REGION Network 108
   RUNG wire#powerrail
      Move(in := "Carrier_05_SDCFaultCode", out1 => "DB_SDC_EMS_TA".EMS[05].TA[1].FAULT)
      wire#w1
      Move(in := "Carrier_05_SDCFaultCode", out1 => "EMS".Carrier[05].SDC_IN.CarrierDriveFaults)
   END_RUNG
   RUNG wire#powerrail
      Contact( "IndiconTempDebugON" )
   END_RUNG wire#w1
   // the same network as SCL:
   "DB_SDC_EMS_TA".EMS[05].TA[1].FAULT := "Carrier_05_SDCFaultCode";
   IF TRUE OR "IndiconTempDebugON" THEN
       "EMS".Carrier[05].SDC_IN.CarrierDriveFaults := "Carrier_05_SDCFaultCode";
   END_IF;
END_REGION

REGION Network 109
   RUNG wire#powerrail
      Move(in := "Carrier_05_CarrierDriveAlarm", out1 => "DB_SDC_EMS_TA".EMS[05].TA[1].ALARM)
      wire#w1
      Move(in := "Carrier_05_CarrierDriveAlarm", out1 => "EMS".Carrier[05].SDC_IN.CarrierDriveAlarms)
   END_RUNG
   RUNG wire#powerrail
      Contact( "IndiconTempDebugON" )
   END_RUNG wire#w1
   // the same network as SCL:
   "DB_SDC_EMS_TA".EMS[05].TA[1].ALARM := "Carrier_05_CarrierDriveAlarm";
   IF TRUE OR "IndiconTempDebugON" THEN
       "EMS".Carrier[05].SDC_IN.CarrierDriveAlarms := "Carrier_05_CarrierDriveAlarm";
   END_IF;
END_REGION

REGION Network 110
   RUNG wire#powerrail
      Move(in := "Carrier_05_SDCFaultCode", out1 => "DB101_DB_SDC_FAULTS".Carrier_Fault[05])
      wire#w1
      Move(in := "Carrier_05_SDCFaultCode", out1 => "EMS".Carrier[05].SDC_IN.CarrierFaults)
   END_RUNG
   RUNG wire#powerrail
      Contact( "IndiconTempDebugON" )
   END_RUNG wire#w1
   // the same network as SCL:
   "DB101_DB_SDC_FAULTS".Carrier_Fault[05] := "Carrier_05_SDCFaultCode";
   IF TRUE OR "IndiconTempDebugON" THEN
       "EMS".Carrier[05].SDC_IN.CarrierFaults := "Carrier_05_SDCFaultCode";
   END_IF;
END_REGION

REGION Network 111
   RUNG wire#powerrail
      Contact( "Carrier_05_Status.5" )
      Coil( "EMS".Carrier[05].SDC_IN.RunningFWD )
   END_RUNG
   // the same network as SCL:
   "EMS".Carrier[05].SDC_IN.RunningFWD := "Carrier_05_Status.5";
END_REGION

REGION Network 112
   RUNG wire#powerrail
      Contact( "Carrier_05_Status.6" )
      Coil( "EMS".Carrier[05].SDC_IN.RunningREV )
   END_RUNG
   // the same network as SCL:
   "EMS".Carrier[05].SDC_IN.RunningREV := "Carrier_05_Status.6";
END_REGION

REGION Network 113
   RUNG wire#powerrail
      Contact( "Carrier_05_Status.7" )
      Coil( "EMS".Carrier[05].SDC_IN.IR_Remote_9_Pressed )
   END_RUNG
   // the same network as SCL:
   "EMS".Carrier[05].SDC_IN.IR_Remote_9_Pressed := "Carrier_05_Status.7";
END_REGION

REGION Network 114
   RUNG wire#powerrail
      I_Contact( "Carrier_05_Status.5" )
      I_Contact( "Carrier_05_Status.6" )
      Coil( "EMS".Carrier[05].SDC_IN.Stopped )
   END_RUNG
   // the same network as SCL:
   "EMS".Carrier[05].SDC_IN.Stopped := NOT "Carrier_05_Status.5" AND NOT "Carrier_05_Status.6";
END_REGION

REGION Network 115
   RUNG wire#powerrail
      Contact( "Carrier_05_Status.4" )
      Coil( "EMS".Carrier[05].SDC_IN.ProductionHoldPB_Status )
   END_RUNG
   // the same network as SCL:
   "EMS".Carrier[05].SDC_IN.ProductionHoldPB_Status := "Carrier_05_Status.4";
END_REGION

REGION Network 116
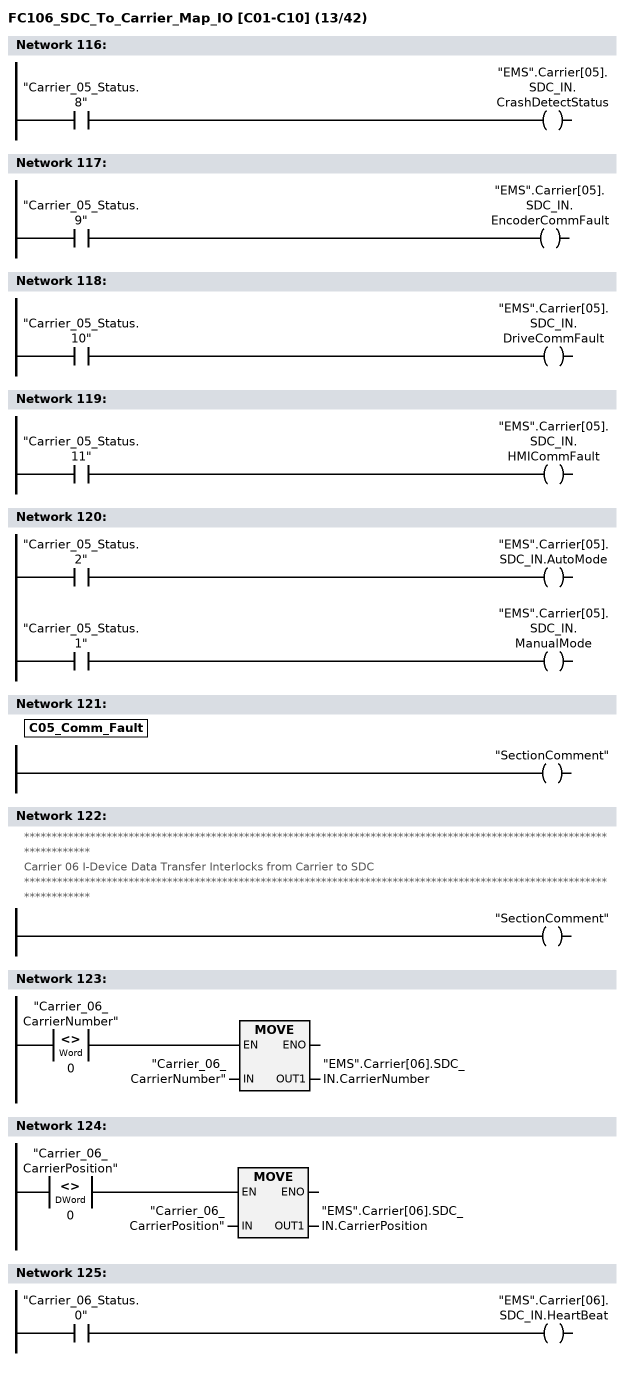
   RUNG wire#powerrail
      Contact( "Carrier_05_Status.8" )
      Coil( "EMS".Carrier[05].SDC_IN.CrashDetectStatus )
   END_RUNG
   // the same network as SCL:
   "EMS".Carrier[05].SDC_IN.CrashDetectStatus := "Carrier_05_Status.8";
END_REGION

REGION Network 117
   RUNG wire#powerrail
      Contact( "Carrier_05_Status.9" )
      Coil( "EMS".Carrier[05].SDC_IN.EncoderCommFault )
   END_RUNG
   // the same network as SCL:
   "EMS".Carrier[05].SDC_IN.EncoderCommFault := "Carrier_05_Status.9";
END_REGION

REGION Network 118
   RUNG wire#powerrail
      Contact( "Carrier_05_Status.10" )
      Coil( "EMS".Carrier[05].SDC_IN.DriveCommFault )
   END_RUNG
   // the same network as SCL:
   "EMS".Carrier[05].SDC_IN.DriveCommFault := "Carrier_05_Status.10";
END_REGION

REGION Network 119
   RUNG wire#powerrail
      Contact( "Carrier_05_Status.11" )
      Coil( "EMS".Carrier[05].SDC_IN.HMICommFault )
   END_RUNG
   // the same network as SCL:
   "EMS".Carrier[05].SDC_IN.HMICommFault := "Carrier_05_Status.11";
END_REGION

REGION Network 120
   RUNG wire#powerrail
      Contact( "Carrier_05_Status.2" )
      Coil( "EMS".Carrier[05].SDC_IN.AutoMode )
   END_RUNG
   RUNG wire#powerrail
      Contact( "Carrier_05_Status.1" )
      Coil( "EMS".Carrier[05].SDC_IN.ManualMode )
   END_RUNG
   // the same network as SCL:
   "EMS".Carrier[05].SDC_IN.AutoMode := "Carrier_05_Status.2";
   "EMS".Carrier[05].SDC_IN.ManualMode := "Carrier_05_Status.1";
END_REGION

REGION Network 121
   Label( C05_Comm_Fault )
   RUNG wire#powerrail
      Coil( "SectionComment" )
   END_RUNG
   // the same network as SCL:
   C05_Comm_Fault:
   "SectionComment" := TRUE;
END_REGION

REGION Network 122
   // **********************************************************************************************************************
   // 
   // Carrier 06 I-Device Data Transfer Interlocks from Carrier to SDC
   // 
   // **********************************************************************************************************************
   RUNG wire#powerrail
      Coil( "SectionComment" )
   END_RUNG
   // the same network as SCL:
   "SectionComment" := TRUE;
END_REGION

REGION Network 123
   RUNG wire#powerrail
      { S7_Templates := "SrcType := Word" } NE_Contact(in1 := "Carrier_06_CarrierNumber", in2 := 0)
      Move(in := "Carrier_06_CarrierNumber", out1 => "EMS".Carrier[06].SDC_IN.CarrierNumber)
   END_RUNG
   // the same network as SCL:
   IF "Carrier_06_CarrierNumber" <> 0 THEN
       "EMS".Carrier[06].SDC_IN.CarrierNumber := "Carrier_06_CarrierNumber";
   END_IF;
END_REGION

REGION Network 124
   RUNG wire#powerrail
      { S7_Templates := "SrcType := DWord" } NE_Contact(in1 := "Carrier_06_CarrierPosition", in2 := 0)
      Move(in := "Carrier_06_CarrierPosition", out1 => "EMS".Carrier[06].SDC_IN.CarrierPosition)
   END_RUNG
   // the same network as SCL:
   IF "Carrier_06_CarrierPosition" <> 0 THEN
       "EMS".Carrier[06].SDC_IN.CarrierPosition := "Carrier_06_CarrierPosition";
   END_IF;
END_REGION

REGION Network 125
   RUNG wire#powerrail
      Contact( "Carrier_06_Status.0" )
      Coil( "EMS".Carrier[06].SDC_IN.HeartBeat )
   END_RUNG
   // the same network as SCL:
   "EMS".Carrier[06].SDC_IN.HeartBeat := "Carrier_06_Status.0";
END_REGION

REGION Network 126
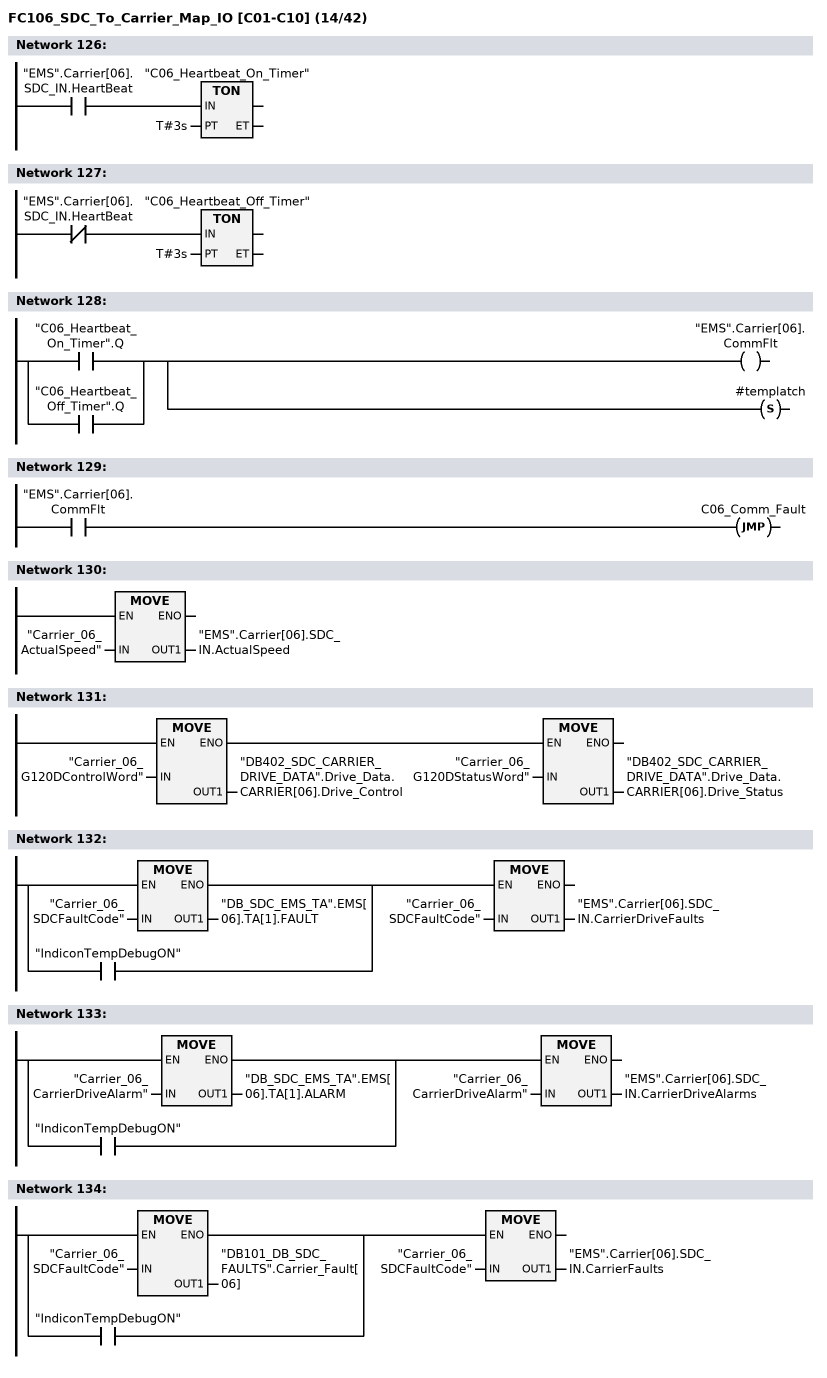
   "C06_Heartbeat_On_Timer".TON(IN := "EMS".Carrier[06].SDC_IN.HeartBeat, PT := T#3s);
END_REGION

REGION Network 127
   "C06_Heartbeat_Off_Timer".TON(IN := NOT "EMS".Carrier[06].SDC_IN.HeartBeat, PT := T#3s);
END_REGION

REGION Network 128
   RUNG wire#powerrail
      Contact( "C06_Heartbeat_On_Timer".Q )
      wire#w1
      Coil( "EMS".Carrier[06].CommFlt )
   END_RUNG
   RUNG wire#powerrail
      Contact( "C06_Heartbeat_Off_Timer".Q )
   END_RUNG wire#w1
   RUNG wire#w1
      S_Coil( #templatch )
   END_RUNG
   // the same network as SCL:
   "EMS".Carrier[06].CommFlt := "C06_Heartbeat_On_Timer".Q OR "C06_Heartbeat_Off_Timer".Q;
   IF "C06_Heartbeat_On_Timer".Q OR "C06_Heartbeat_Off_Timer".Q THEN #templatch := TRUE; END_IF;
END_REGION

REGION Network 129
   RUNG wire#powerrail
      Contact( "EMS".Carrier[06].CommFlt )
      JumpCoil( C06_Comm_Fault )
   END_RUNG
   // the same network as SCL:
   IF "EMS".Carrier[06].CommFlt THEN GOTO C06_Comm_Fault; END_IF;
END_REGION

REGION Network 130
   RUNG wire#powerrail
      Move(in := "Carrier_06_ActualSpeed", out1 => "EMS".Carrier[06].SDC_IN.ActualSpeed)
   END_RUNG
   // the same network as SCL:
   "EMS".Carrier[06].SDC_IN.ActualSpeed := "Carrier_06_ActualSpeed";
END_REGION

REGION Network 131
   RUNG wire#powerrail
      Move(in := "Carrier_06_G120DControlWord", out1 => "DB402_SDC_CARRIER_DRIVE_DATA".Drive_Data.CARRIER[06].Drive_Control)
      Move(in := "Carrier_06_G120DStatusWord", out1 => "DB402_SDC_CARRIER_DRIVE_DATA".Drive_Data.CARRIER[06].Drive_Status)
   END_RUNG
   // the same network as SCL:
   "DB402_SDC_CARRIER_DRIVE_DATA".Drive_Data.CARRIER[06].Drive_Control := "Carrier_06_G120DControlWord";
   "DB402_SDC_CARRIER_DRIVE_DATA".Drive_Data.CARRIER[06].Drive_Status := "Carrier_06_G120DStatusWord";
END_REGION

REGION Network 132
   RUNG wire#powerrail
      Move(in := "Carrier_06_SDCFaultCode", out1 => "DB_SDC_EMS_TA".EMS[06].TA[1].FAULT)
      wire#w1
      Move(in := "Carrier_06_SDCFaultCode", out1 => "EMS".Carrier[06].SDC_IN.CarrierDriveFaults)
   END_RUNG
   RUNG wire#powerrail
      Contact( "IndiconTempDebugON" )
   END_RUNG wire#w1
   // the same network as SCL:
   "DB_SDC_EMS_TA".EMS[06].TA[1].FAULT := "Carrier_06_SDCFaultCode";
   IF TRUE OR "IndiconTempDebugON" THEN
       "EMS".Carrier[06].SDC_IN.CarrierDriveFaults := "Carrier_06_SDCFaultCode";
   END_IF;
END_REGION

REGION Network 133
   RUNG wire#powerrail
      Move(in := "Carrier_06_CarrierDriveAlarm", out1 => "DB_SDC_EMS_TA".EMS[06].TA[1].ALARM)
      wire#w1
      Move(in := "Carrier_06_CarrierDriveAlarm", out1 => "EMS".Carrier[06].SDC_IN.CarrierDriveAlarms)
   END_RUNG
   RUNG wire#powerrail
      Contact( "IndiconTempDebugON" )
   END_RUNG wire#w1
   // the same network as SCL:
   "DB_SDC_EMS_TA".EMS[06].TA[1].ALARM := "Carrier_06_CarrierDriveAlarm";
   IF TRUE OR "IndiconTempDebugON" THEN
       "EMS".Carrier[06].SDC_IN.CarrierDriveAlarms := "Carrier_06_CarrierDriveAlarm";
   END_IF;
END_REGION

REGION Network 134
   RUNG wire#powerrail
      Move(in := "Carrier_06_SDCFaultCode", out1 => "DB101_DB_SDC_FAULTS".Carrier_Fault[06])
      wire#w1
      Move(in := "Carrier_06_SDCFaultCode", out1 => "EMS".Carrier[06].SDC_IN.CarrierFaults)
   END_RUNG
   RUNG wire#powerrail
      Contact( "IndiconTempDebugON" )
   END_RUNG wire#w1
   // the same network as SCL:
   "DB101_DB_SDC_FAULTS".Carrier_Fault[06] := "Carrier_06_SDCFaultCode";
   IF TRUE OR "IndiconTempDebugON" THEN
       "EMS".Carrier[06].SDC_IN.CarrierFaults := "Carrier_06_SDCFaultCode";
   END_IF;
END_REGION

REGION Network 135
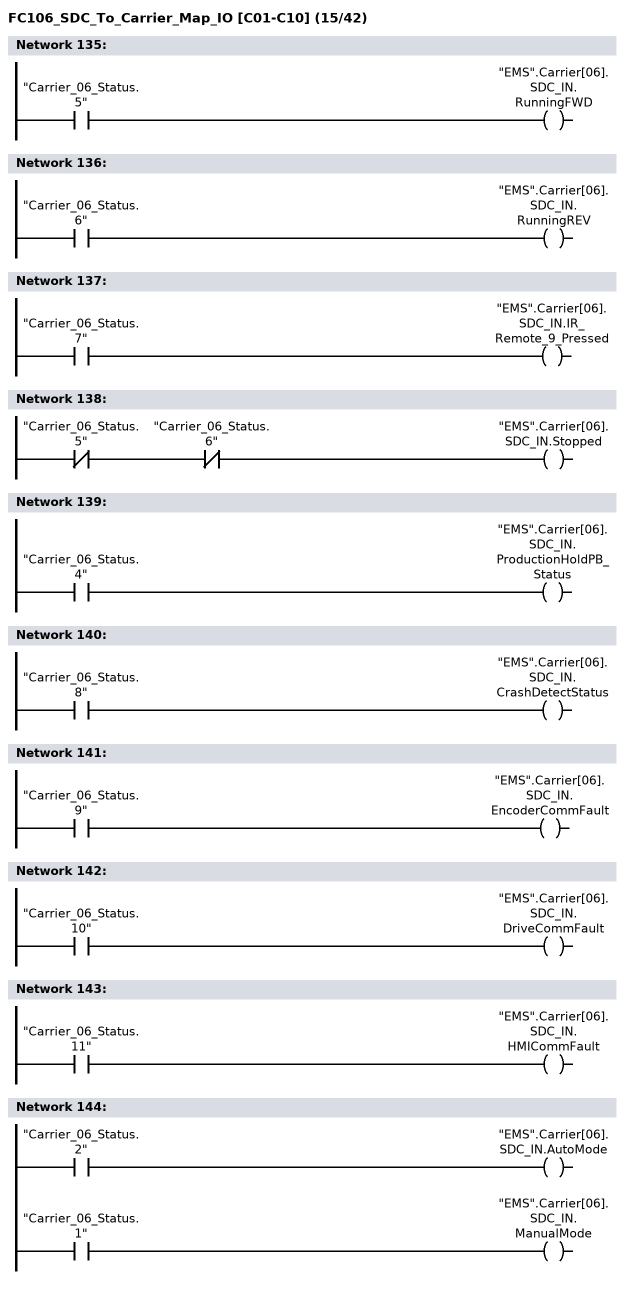
   RUNG wire#powerrail
      Contact( "Carrier_06_Status.5" )
      Coil( "EMS".Carrier[06].SDC_IN.RunningFWD )
   END_RUNG
   // the same network as SCL:
   "EMS".Carrier[06].SDC_IN.RunningFWD := "Carrier_06_Status.5";
END_REGION

REGION Network 136
   RUNG wire#powerrail
      Contact( "Carrier_06_Status.6" )
      Coil( "EMS".Carrier[06].SDC_IN.RunningREV )
   END_RUNG
   // the same network as SCL:
   "EMS".Carrier[06].SDC_IN.RunningREV := "Carrier_06_Status.6";
END_REGION

REGION Network 137
   RUNG wire#powerrail
      Contact( "Carrier_06_Status.7" )
      Coil( "EMS".Carrier[06].SDC_IN.IR_Remote_9_Pressed )
   END_RUNG
   // the same network as SCL:
   "EMS".Carrier[06].SDC_IN.IR_Remote_9_Pressed := "Carrier_06_Status.7";
END_REGION

REGION Network 138
   RUNG wire#powerrail
      I_Contact( "Carrier_06_Status.5" )
      I_Contact( "Carrier_06_Status.6" )
      Coil( "EMS".Carrier[06].SDC_IN.Stopped )
   END_RUNG
   // the same network as SCL:
   "EMS".Carrier[06].SDC_IN.Stopped := NOT "Carrier_06_Status.5" AND NOT "Carrier_06_Status.6";
END_REGION

REGION Network 139
   RUNG wire#powerrail
      Contact( "Carrier_06_Status.4" )
      Coil( "EMS".Carrier[06].SDC_IN.ProductionHoldPB_Status )
   END_RUNG
   // the same network as SCL:
   "EMS".Carrier[06].SDC_IN.ProductionHoldPB_Status := "Carrier_06_Status.4";
END_REGION

REGION Network 140
   RUNG wire#powerrail
      Contact( "Carrier_06_Status.8" )
      Coil( "EMS".Carrier[06].SDC_IN.CrashDetectStatus )
   END_RUNG
   // the same network as SCL:
   "EMS".Carrier[06].SDC_IN.CrashDetectStatus := "Carrier_06_Status.8";
END_REGION

REGION Network 141
   RUNG wire#powerrail
      Contact( "Carrier_06_Status.9" )
      Coil( "EMS".Carrier[06].SDC_IN.EncoderCommFault )
   END_RUNG
   // the same network as SCL:
   "EMS".Carrier[06].SDC_IN.EncoderCommFault := "Carrier_06_Status.9";
END_REGION

REGION Network 142
   RUNG wire#powerrail
      Contact( "Carrier_06_Status.10" )
      Coil( "EMS".Carrier[06].SDC_IN.DriveCommFault )
   END_RUNG
   // the same network as SCL:
   "EMS".Carrier[06].SDC_IN.DriveCommFault := "Carrier_06_Status.10";
END_REGION

REGION Network 143
   RUNG wire#powerrail
      Contact( "Carrier_06_Status.11" )
      Coil( "EMS".Carrier[06].SDC_IN.HMICommFault )
   END_RUNG
   // the same network as SCL:
   "EMS".Carrier[06].SDC_IN.HMICommFault := "Carrier_06_Status.11";
END_REGION

REGION Network 144
   RUNG wire#powerrail
      Contact( "Carrier_06_Status.2" )
      Coil( "EMS".Carrier[06].SDC_IN.AutoMode )
   END_RUNG
   RUNG wire#powerrail
      Contact( "Carrier_06_Status.1" )
      Coil( "EMS".Carrier[06].SDC_IN.ManualMode )
   END_RUNG
   // the same network as SCL:
   "EMS".Carrier[06].SDC_IN.AutoMode := "Carrier_06_Status.2";
   "EMS".Carrier[06].SDC_IN.ManualMode := "Carrier_06_Status.1";
END_REGION

REGION Network 145
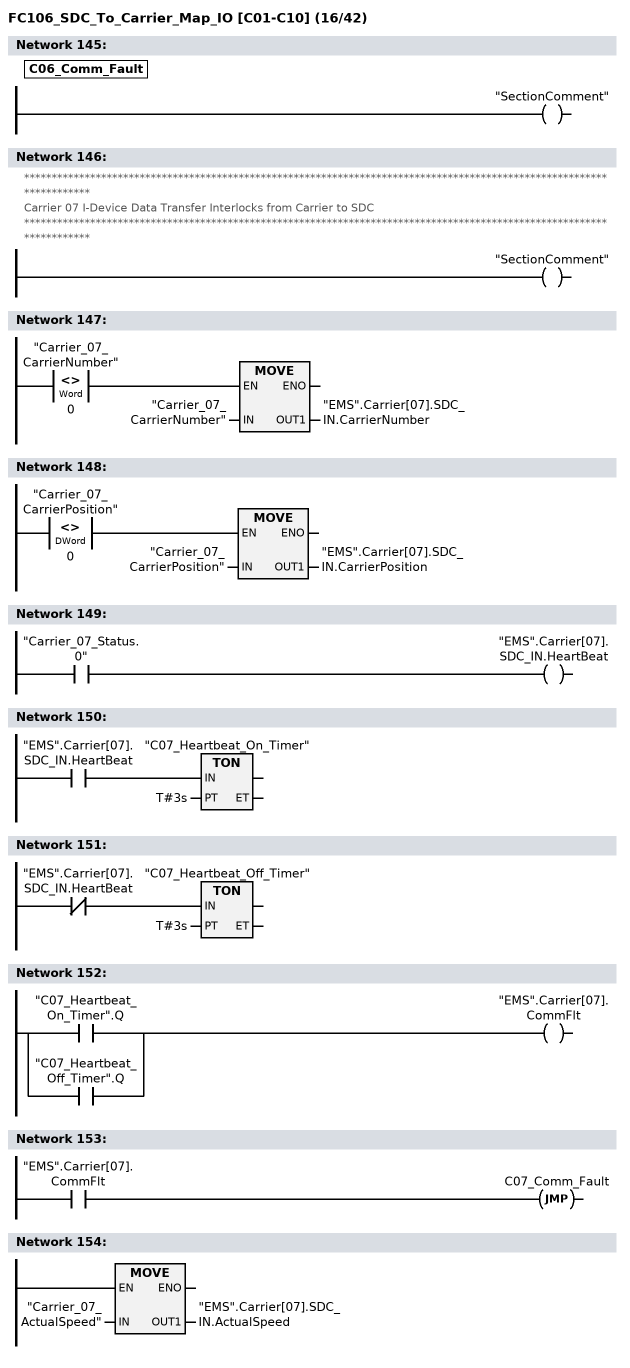
   Label( C06_Comm_Fault )
   RUNG wire#powerrail
      Coil( "SectionComment" )
   END_RUNG
   // the same network as SCL:
   C06_Comm_Fault:
   "SectionComment" := TRUE;
END_REGION

REGION Network 146
   // **********************************************************************************************************************
   // 
   // Carrier 07 I-Device Data Transfer Interlocks from Carrier to SDC
   // 
   // **********************************************************************************************************************
   RUNG wire#powerrail
      Coil( "SectionComment" )
   END_RUNG
   // the same network as SCL:
   "SectionComment" := TRUE;
END_REGION

REGION Network 147
   RUNG wire#powerrail
      { S7_Templates := "SrcType := Word" } NE_Contact(in1 := "Carrier_07_CarrierNumber", in2 := 0)
      Move(in := "Carrier_07_CarrierNumber", out1 => "EMS".Carrier[07].SDC_IN.CarrierNumber)
   END_RUNG
   // the same network as SCL:
   IF "Carrier_07_CarrierNumber" <> 0 THEN
       "EMS".Carrier[07].SDC_IN.CarrierNumber := "Carrier_07_CarrierNumber";
   END_IF;
END_REGION

REGION Network 148
   RUNG wire#powerrail
      { S7_Templates := "SrcType := DWord" } NE_Contact(in1 := "Carrier_07_CarrierPosition", in2 := 0)
      Move(in := "Carrier_07_CarrierPosition", out1 => "EMS".Carrier[07].SDC_IN.CarrierPosition)
   END_RUNG
   // the same network as SCL:
   IF "Carrier_07_CarrierPosition" <> 0 THEN
       "EMS".Carrier[07].SDC_IN.CarrierPosition := "Carrier_07_CarrierPosition";
   END_IF;
END_REGION

REGION Network 149
   RUNG wire#powerrail
      Contact( "Carrier_07_Status.0" )
      Coil( "EMS".Carrier[07].SDC_IN.HeartBeat )
   END_RUNG
   // the same network as SCL:
   "EMS".Carrier[07].SDC_IN.HeartBeat := "Carrier_07_Status.0";
END_REGION

REGION Network 150
   "C07_Heartbeat_On_Timer".TON(IN := "EMS".Carrier[07].SDC_IN.HeartBeat, PT := T#3s);
END_REGION

REGION Network 151
   "C07_Heartbeat_Off_Timer".TON(IN := NOT "EMS".Carrier[07].SDC_IN.HeartBeat, PT := T#3s);
END_REGION

REGION Network 152
   RUNG wire#powerrail
      Contact( "C07_Heartbeat_On_Timer".Q )
      wire#w1
      Coil( "EMS".Carrier[07].CommFlt )
   END_RUNG
   RUNG wire#powerrail
      Contact( "C07_Heartbeat_Off_Timer".Q )
   END_RUNG wire#w1
   // the same network as SCL:
   "EMS".Carrier[07].CommFlt := "C07_Heartbeat_On_Timer".Q OR "C07_Heartbeat_Off_Timer".Q;
END_REGION

REGION Network 153
   RUNG wire#powerrail
      Contact( "EMS".Carrier[07].CommFlt )
      JumpCoil( C07_Comm_Fault )
   END_RUNG
   // the same network as SCL:
   IF "EMS".Carrier[07].CommFlt THEN GOTO C07_Comm_Fault; END_IF;
END_REGION

REGION Network 154
   RUNG wire#powerrail
      Move(in := "Carrier_07_ActualSpeed", out1 => "EMS".Carrier[07].SDC_IN.ActualSpeed)
   END_RUNG
   // the same network as SCL:
   "EMS".Carrier[07].SDC_IN.ActualSpeed := "Carrier_07_ActualSpeed";
END_REGION

REGION Network 155
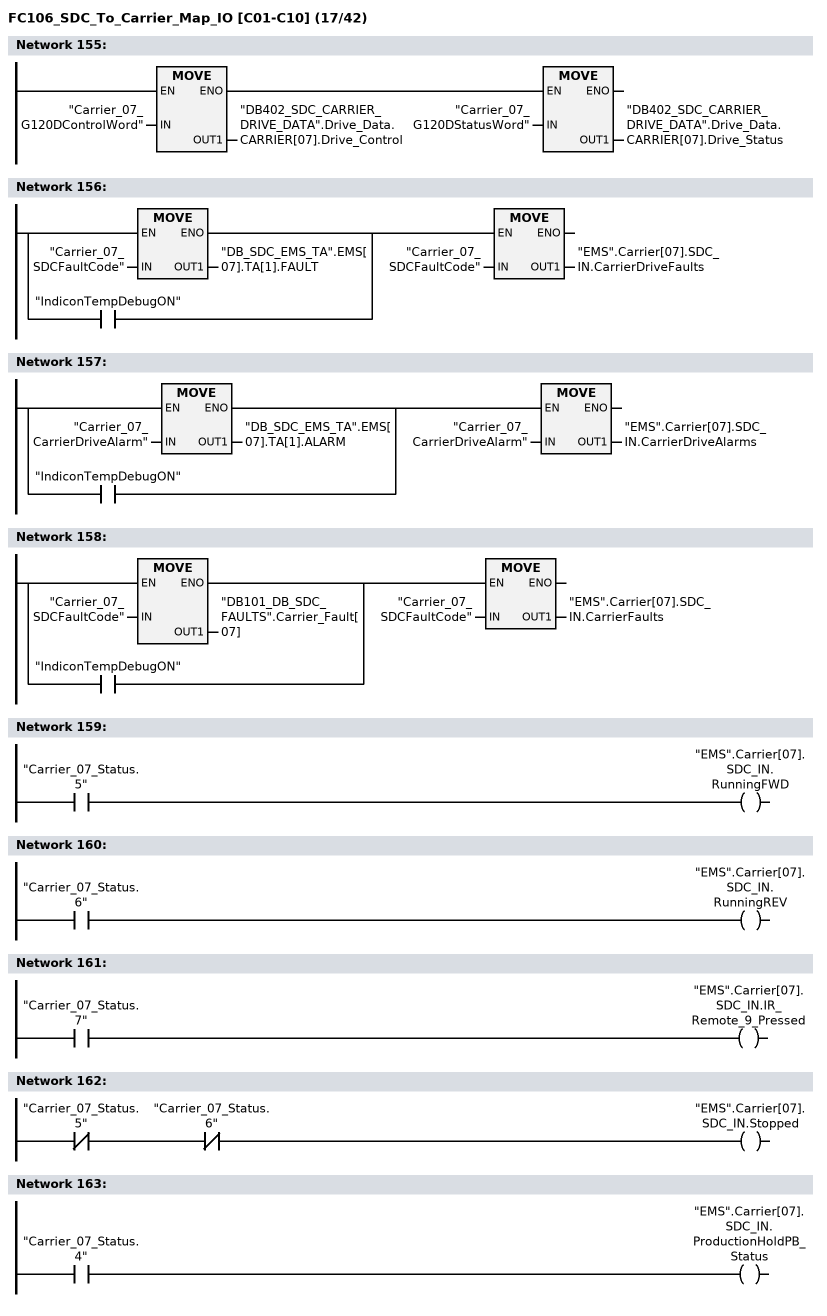
   RUNG wire#powerrail
      Move(in := "Carrier_07_G120DControlWord", out1 => "DB402_SDC_CARRIER_DRIVE_DATA".Drive_Data.CARRIER[07].Drive_Control)
      Move(in := "Carrier_07_G120DStatusWord", out1 => "DB402_SDC_CARRIER_DRIVE_DATA".Drive_Data.CARRIER[07].Drive_Status)
   END_RUNG
   // the same network as SCL:
   "DB402_SDC_CARRIER_DRIVE_DATA".Drive_Data.CARRIER[07].Drive_Control := "Carrier_07_G120DControlWord";
   "DB402_SDC_CARRIER_DRIVE_DATA".Drive_Data.CARRIER[07].Drive_Status := "Carrier_07_G120DStatusWord";
END_REGION

REGION Network 156
   RUNG wire#powerrail
      Move(in := "Carrier_07_SDCFaultCode", out1 => "DB_SDC_EMS_TA".EMS[07].TA[1].FAULT)
      wire#w1
      Move(in := "Carrier_07_SDCFaultCode", out1 => "EMS".Carrier[07].SDC_IN.CarrierDriveFaults)
   END_RUNG
   RUNG wire#powerrail
      Contact( "IndiconTempDebugON" )
   END_RUNG wire#w1
   // the same network as SCL:
   "DB_SDC_EMS_TA".EMS[07].TA[1].FAULT := "Carrier_07_SDCFaultCode";
   IF TRUE OR "IndiconTempDebugON" THEN
       "EMS".Carrier[07].SDC_IN.CarrierDriveFaults := "Carrier_07_SDCFaultCode";
   END_IF;
END_REGION

REGION Network 157
   RUNG wire#powerrail
      Move(in := "Carrier_07_CarrierDriveAlarm", out1 => "DB_SDC_EMS_TA".EMS[07].TA[1].ALARM)
      wire#w1
      Move(in := "Carrier_07_CarrierDriveAlarm", out1 => "EMS".Carrier[07].SDC_IN.CarrierDriveAlarms)
   END_RUNG
   RUNG wire#powerrail
      Contact( "IndiconTempDebugON" )
   END_RUNG wire#w1
   // the same network as SCL:
   "DB_SDC_EMS_TA".EMS[07].TA[1].ALARM := "Carrier_07_CarrierDriveAlarm";
   IF TRUE OR "IndiconTempDebugON" THEN
       "EMS".Carrier[07].SDC_IN.CarrierDriveAlarms := "Carrier_07_CarrierDriveAlarm";
   END_IF;
END_REGION

REGION Network 158
   RUNG wire#powerrail
      Move(in := "Carrier_07_SDCFaultCode", out1 => "DB101_DB_SDC_FAULTS".Carrier_Fault[07])
      wire#w1
      Move(in := "Carrier_07_SDCFaultCode", out1 => "EMS".Carrier[07].SDC_IN.CarrierFaults)
   END_RUNG
   RUNG wire#powerrail
      Contact( "IndiconTempDebugON" )
   END_RUNG wire#w1
   // the same network as SCL:
   "DB101_DB_SDC_FAULTS".Carrier_Fault[07] := "Carrier_07_SDCFaultCode";
   IF TRUE OR "IndiconTempDebugON" THEN
       "EMS".Carrier[07].SDC_IN.CarrierFaults := "Carrier_07_SDCFaultCode";
   END_IF;
END_REGION

REGION Network 159
   RUNG wire#powerrail
      Contact( "Carrier_07_Status.5" )
      Coil( "EMS".Carrier[07].SDC_IN.RunningFWD )
   END_RUNG
   // the same network as SCL:
   "EMS".Carrier[07].SDC_IN.RunningFWD := "Carrier_07_Status.5";
END_REGION

REGION Network 160
   RUNG wire#powerrail
      Contact( "Carrier_07_Status.6" )
      Coil( "EMS".Carrier[07].SDC_IN.RunningREV )
   END_RUNG
   // the same network as SCL:
   "EMS".Carrier[07].SDC_IN.RunningREV := "Carrier_07_Status.6";
END_REGION

REGION Network 161
   RUNG wire#powerrail
      Contact( "Carrier_07_Status.7" )
      Coil( "EMS".Carrier[07].SDC_IN.IR_Remote_9_Pressed )
   END_RUNG
   // the same network as SCL:
   "EMS".Carrier[07].SDC_IN.IR_Remote_9_Pressed := "Carrier_07_Status.7";
END_REGION

REGION Network 162
   RUNG wire#powerrail
      I_Contact( "Carrier_07_Status.5" )
      I_Contact( "Carrier_07_Status.6" )
      Coil( "EMS".Carrier[07].SDC_IN.Stopped )
   END_RUNG
   // the same network as SCL:
   "EMS".Carrier[07].SDC_IN.Stopped := NOT "Carrier_07_Status.5" AND NOT "Carrier_07_Status.6";
END_REGION

REGION Network 163
   RUNG wire#powerrail
      Contact( "Carrier_07_Status.4" )
      Coil( "EMS".Carrier[07].SDC_IN.ProductionHoldPB_Status )
   END_RUNG
   // the same network as SCL:
   "EMS".Carrier[07].SDC_IN.ProductionHoldPB_Status := "Carrier_07_Status.4";
END_REGION

REGION Network 164
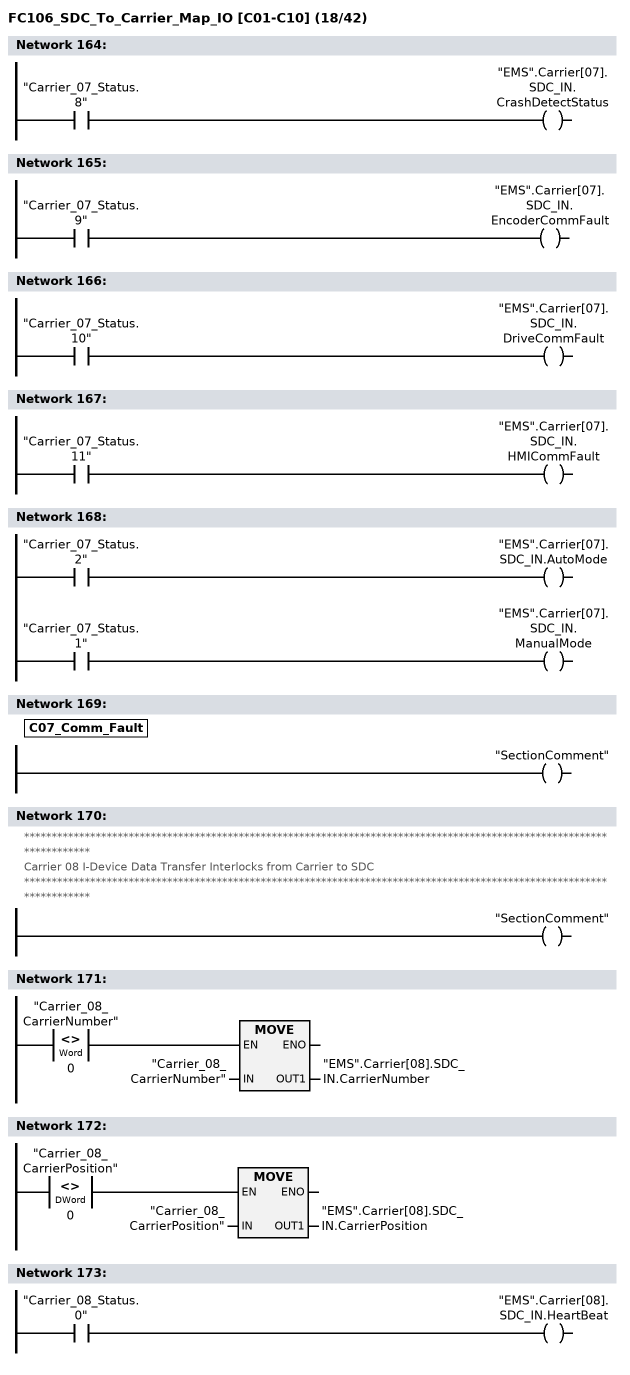
   RUNG wire#powerrail
      Contact( "Carrier_07_Status.8" )
      Coil( "EMS".Carrier[07].SDC_IN.CrashDetectStatus )
   END_RUNG
   // the same network as SCL:
   "EMS".Carrier[07].SDC_IN.CrashDetectStatus := "Carrier_07_Status.8";
END_REGION

REGION Network 165
   RUNG wire#powerrail
      Contact( "Carrier_07_Status.9" )
      Coil( "EMS".Carrier[07].SDC_IN.EncoderCommFault )
   END_RUNG
   // the same network as SCL:
   "EMS".Carrier[07].SDC_IN.EncoderCommFault := "Carrier_07_Status.9";
END_REGION

REGION Network 166
   RUNG wire#powerrail
      Contact( "Carrier_07_Status.10" )
      Coil( "EMS".Carrier[07].SDC_IN.DriveCommFault )
   END_RUNG
   // the same network as SCL:
   "EMS".Carrier[07].SDC_IN.DriveCommFault := "Carrier_07_Status.10";
END_REGION

REGION Network 167
   RUNG wire#powerrail
      Contact( "Carrier_07_Status.11" )
      Coil( "EMS".Carrier[07].SDC_IN.HMICommFault )
   END_RUNG
   // the same network as SCL:
   "EMS".Carrier[07].SDC_IN.HMICommFault := "Carrier_07_Status.11";
END_REGION

REGION Network 168
   RUNG wire#powerrail
      Contact( "Carrier_07_Status.2" )
      Coil( "EMS".Carrier[07].SDC_IN.AutoMode )
   END_RUNG
   RUNG wire#powerrail
      Contact( "Carrier_07_Status.1" )
      Coil( "EMS".Carrier[07].SDC_IN.ManualMode )
   END_RUNG
   // the same network as SCL:
   "EMS".Carrier[07].SDC_IN.AutoMode := "Carrier_07_Status.2";
   "EMS".Carrier[07].SDC_IN.ManualMode := "Carrier_07_Status.1";
END_REGION

REGION Network 169
   Label( C07_Comm_Fault )
   RUNG wire#powerrail
      Coil( "SectionComment" )
   END_RUNG
   // the same network as SCL:
   C07_Comm_Fault:
   "SectionComment" := TRUE;
END_REGION

REGION Network 170
   // **********************************************************************************************************************
   // 
   // Carrier 08 I-Device Data Transfer Interlocks from Carrier to SDC
   // 
   // **********************************************************************************************************************
   RUNG wire#powerrail
      Coil( "SectionComment" )
   END_RUNG
   // the same network as SCL:
   "SectionComment" := TRUE;
END_REGION

REGION Network 171
   RUNG wire#powerrail
      { S7_Templates := "SrcType := Word" } NE_Contact(in1 := "Carrier_08_CarrierNumber", in2 := 0)
      Move(in := "Carrier_08_CarrierNumber", out1 => "EMS".Carrier[08].SDC_IN.CarrierNumber)
   END_RUNG
   // the same network as SCL:
   IF "Carrier_08_CarrierNumber" <> 0 THEN
       "EMS".Carrier[08].SDC_IN.CarrierNumber := "Carrier_08_CarrierNumber";
   END_IF;
END_REGION

REGION Network 172
   RUNG wire#powerrail
      { S7_Templates := "SrcType := DWord" } NE_Contact(in1 := "Carrier_08_CarrierPosition", in2 := 0)
      Move(in := "Carrier_08_CarrierPosition", out1 => "EMS".Carrier[08].SDC_IN.CarrierPosition)
   END_RUNG
   // the same network as SCL:
   IF "Carrier_08_CarrierPosition" <> 0 THEN
       "EMS".Carrier[08].SDC_IN.CarrierPosition := "Carrier_08_CarrierPosition";
   END_IF;
END_REGION

REGION Network 173
   RUNG wire#powerrail
      Contact( "Carrier_08_Status.0" )
      Coil( "EMS".Carrier[08].SDC_IN.HeartBeat )
   END_RUNG
   // the same network as SCL:
   "EMS".Carrier[08].SDC_IN.HeartBeat := "Carrier_08_Status.0";
END_REGION

REGION Network 174
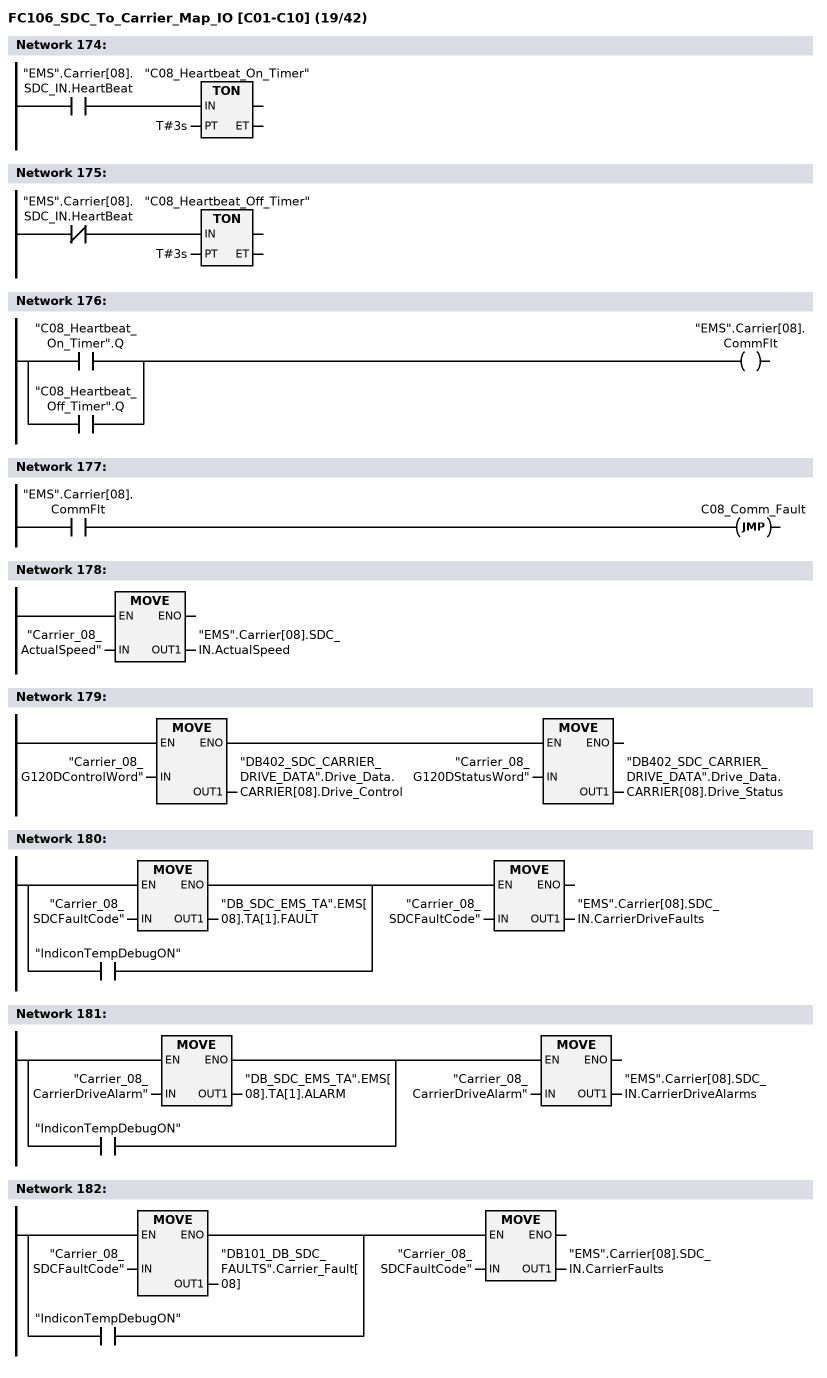
   "C08_Heartbeat_On_Timer".TON(IN := "EMS".Carrier[08].SDC_IN.HeartBeat, PT := T#3s);
END_REGION

REGION Network 175
   "C08_Heartbeat_Off_Timer".TON(IN := NOT "EMS".Carrier[08].SDC_IN.HeartBeat, PT := T#3s);
END_REGION

REGION Network 176
   RUNG wire#powerrail
      Contact( "C08_Heartbeat_On_Timer".Q )
      wire#w1
      Coil( "EMS".Carrier[08].CommFlt )
   END_RUNG
   RUNG wire#powerrail
      Contact( "C08_Heartbeat_Off_Timer".Q )
   END_RUNG wire#w1
   // the same network as SCL:
   "EMS".Carrier[08].CommFlt := "C08_Heartbeat_On_Timer".Q OR "C08_Heartbeat_Off_Timer".Q;
END_REGION

REGION Network 177
   RUNG wire#powerrail
      Contact( "EMS".Carrier[08].CommFlt )
      JumpCoil( C08_Comm_Fault )
   END_RUNG
   // the same network as SCL:
   IF "EMS".Carrier[08].CommFlt THEN GOTO C08_Comm_Fault; END_IF;
END_REGION

REGION Network 178
   RUNG wire#powerrail
      Move(in := "Carrier_08_ActualSpeed", out1 => "EMS".Carrier[08].SDC_IN.ActualSpeed)
   END_RUNG
   // the same network as SCL:
   "EMS".Carrier[08].SDC_IN.ActualSpeed := "Carrier_08_ActualSpeed";
END_REGION

REGION Network 179
   RUNG wire#powerrail
      Move(in := "Carrier_08_G120DControlWord", out1 => "DB402_SDC_CARRIER_DRIVE_DATA".Drive_Data.CARRIER[08].Drive_Control)
      Move(in := "Carrier_08_G120DStatusWord", out1 => "DB402_SDC_CARRIER_DRIVE_DATA".Drive_Data.CARRIER[08].Drive_Status)
   END_RUNG
   // the same network as SCL:
   "DB402_SDC_CARRIER_DRIVE_DATA".Drive_Data.CARRIER[08].Drive_Control := "Carrier_08_G120DControlWord";
   "DB402_SDC_CARRIER_DRIVE_DATA".Drive_Data.CARRIER[08].Drive_Status := "Carrier_08_G120DStatusWord";
END_REGION

REGION Network 180
   RUNG wire#powerrail
      Move(in := "Carrier_08_SDCFaultCode", out1 => "DB_SDC_EMS_TA".EMS[08].TA[1].FAULT)
      wire#w1
      Move(in := "Carrier_08_SDCFaultCode", out1 => "EMS".Carrier[08].SDC_IN.CarrierDriveFaults)
   END_RUNG
   RUNG wire#powerrail
      Contact( "IndiconTempDebugON" )
   END_RUNG wire#w1
   // the same network as SCL:
   "DB_SDC_EMS_TA".EMS[08].TA[1].FAULT := "Carrier_08_SDCFaultCode";
   IF TRUE OR "IndiconTempDebugON" THEN
       "EMS".Carrier[08].SDC_IN.CarrierDriveFaults := "Carrier_08_SDCFaultCode";
   END_IF;
END_REGION

REGION Network 181
   RUNG wire#powerrail
      Move(in := "Carrier_08_CarrierDriveAlarm", out1 => "DB_SDC_EMS_TA".EMS[08].TA[1].ALARM)
      wire#w1
      Move(in := "Carrier_08_CarrierDriveAlarm", out1 => "EMS".Carrier[08].SDC_IN.CarrierDriveAlarms)
   END_RUNG
   RUNG wire#powerrail
      Contact( "IndiconTempDebugON" )
   END_RUNG wire#w1
   // the same network as SCL:
   "DB_SDC_EMS_TA".EMS[08].TA[1].ALARM := "Carrier_08_CarrierDriveAlarm";
   IF TRUE OR "IndiconTempDebugON" THEN
       "EMS".Carrier[08].SDC_IN.CarrierDriveAlarms := "Carrier_08_CarrierDriveAlarm";
   END_IF;
END_REGION

REGION Network 182
   RUNG wire#powerrail
      Move(in := "Carrier_08_SDCFaultCode", out1 => "DB101_DB_SDC_FAULTS".Carrier_Fault[08])
      wire#w1
      Move(in := "Carrier_08_SDCFaultCode", out1 => "EMS".Carrier[08].SDC_IN.CarrierFaults)
   END_RUNG
   RUNG wire#powerrail
      Contact( "IndiconTempDebugON" )
   END_RUNG wire#w1
   // the same network as SCL:
   "DB101_DB_SDC_FAULTS".Carrier_Fault[08] := "Carrier_08_SDCFaultCode";
   IF TRUE OR "IndiconTempDebugON" THEN
       "EMS".Carrier[08].SDC_IN.CarrierFaults := "Carrier_08_SDCFaultCode";
   END_IF;
END_REGION

REGION Network 183
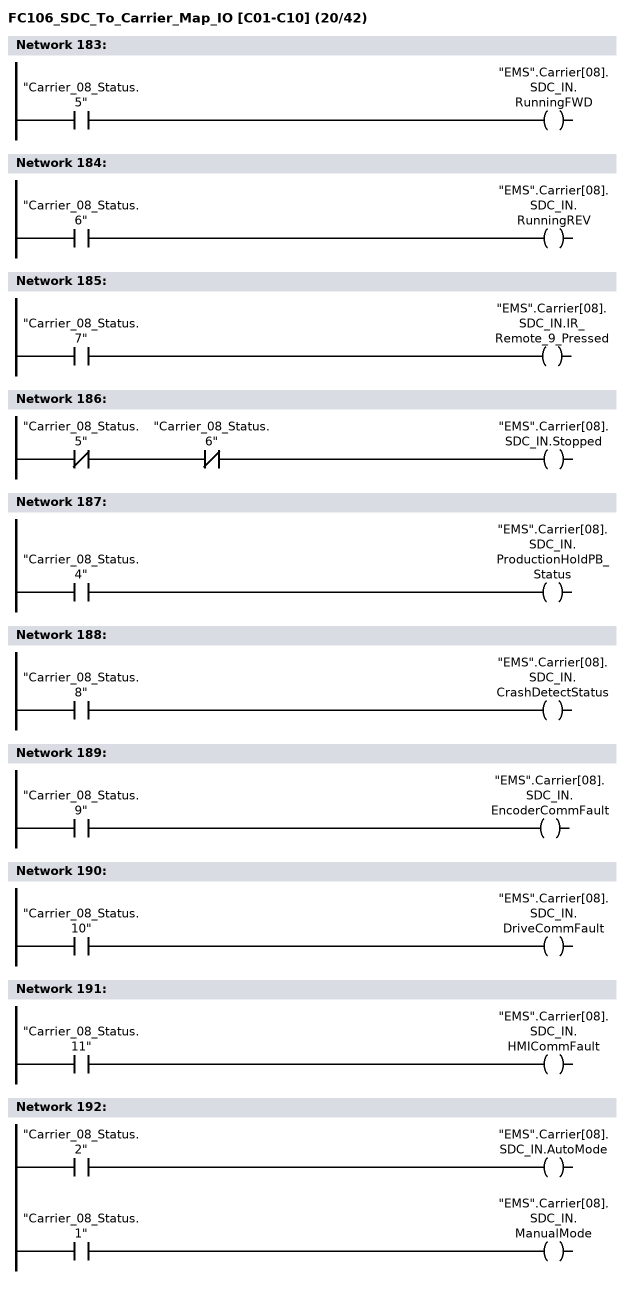
   RUNG wire#powerrail
      Contact( "Carrier_08_Status.5" )
      Coil( "EMS".Carrier[08].SDC_IN.RunningFWD )
   END_RUNG
   // the same network as SCL:
   "EMS".Carrier[08].SDC_IN.RunningFWD := "Carrier_08_Status.5";
END_REGION

REGION Network 184
   RUNG wire#powerrail
      Contact( "Carrier_08_Status.6" )
      Coil( "EMS".Carrier[08].SDC_IN.RunningREV )
   END_RUNG
   // the same network as SCL:
   "EMS".Carrier[08].SDC_IN.RunningREV := "Carrier_08_Status.6";
END_REGION

REGION Network 185
   RUNG wire#powerrail
      Contact( "Carrier_08_Status.7" )
      Coil( "EMS".Carrier[08].SDC_IN.IR_Remote_9_Pressed )
   END_RUNG
   // the same network as SCL:
   "EMS".Carrier[08].SDC_IN.IR_Remote_9_Pressed := "Carrier_08_Status.7";
END_REGION

REGION Network 186
   RUNG wire#powerrail
      I_Contact( "Carrier_08_Status.5" )
      I_Contact( "Carrier_08_Status.6" )
      Coil( "EMS".Carrier[08].SDC_IN.Stopped )
   END_RUNG
   // the same network as SCL:
   "EMS".Carrier[08].SDC_IN.Stopped := NOT "Carrier_08_Status.5" AND NOT "Carrier_08_Status.6";
END_REGION

REGION Network 187
   RUNG wire#powerrail
      Contact( "Carrier_08_Status.4" )
      Coil( "EMS".Carrier[08].SDC_IN.ProductionHoldPB_Status )
   END_RUNG
   // the same network as SCL:
   "EMS".Carrier[08].SDC_IN.ProductionHoldPB_Status := "Carrier_08_Status.4";
END_REGION

REGION Network 188
   RUNG wire#powerrail
      Contact( "Carrier_08_Status.8" )
      Coil( "EMS".Carrier[08].SDC_IN.CrashDetectStatus )
   END_RUNG
   // the same network as SCL:
   "EMS".Carrier[08].SDC_IN.CrashDetectStatus := "Carrier_08_Status.8";
END_REGION

REGION Network 189
   RUNG wire#powerrail
      Contact( "Carrier_08_Status.9" )
      Coil( "EMS".Carrier[08].SDC_IN.EncoderCommFault )
   END_RUNG
   // the same network as SCL:
   "EMS".Carrier[08].SDC_IN.EncoderCommFault := "Carrier_08_Status.9";
END_REGION

REGION Network 190
   RUNG wire#powerrail
      Contact( "Carrier_08_Status.10" )
      Coil( "EMS".Carrier[08].SDC_IN.DriveCommFault )
   END_RUNG
   // the same network as SCL:
   "EMS".Carrier[08].SDC_IN.DriveCommFault := "Carrier_08_Status.10";
END_REGION

REGION Network 191
   RUNG wire#powerrail
      Contact( "Carrier_08_Status.11" )
      Coil( "EMS".Carrier[08].SDC_IN.HMICommFault )
   END_RUNG
   // the same network as SCL:
   "EMS".Carrier[08].SDC_IN.HMICommFault := "Carrier_08_Status.11";
END_REGION

REGION Network 192
   RUNG wire#powerrail
      Contact( "Carrier_08_Status.2" )
      Coil( "EMS".Carrier[08].SDC_IN.AutoMode )
   END_RUNG
   RUNG wire#powerrail
      Contact( "Carrier_08_Status.1" )
      Coil( "EMS".Carrier[08].SDC_IN.ManualMode )
   END_RUNG
   // the same network as SCL:
   "EMS".Carrier[08].SDC_IN.AutoMode := "Carrier_08_Status.2";
   "EMS".Carrier[08].SDC_IN.ManualMode := "Carrier_08_Status.1";
END_REGION

REGION Network 193
